// TIA Portal project "Inteligenta_szklarnia" (V15.1)

(* hardware
DEVICE "S7-1200 station_2"  S7-1200 Station
   slot 0: "Rack_0"  S7-1200 Rack  Rack  V1.0
   slot 1: "PLC_1"  CPU 1214C AC/DC/Rly  6ES7 214-1BE30-0XB0  V2.2
DEVICE "HMI_1"  KTP700 Basic PN
   slot 0: "HMI_1"  KTP700 Basic PN  6AV2 123-2GB03-0AX0  15.1.0.0
   slot 1: "HMI_RT_3"  KTP700 Basic PN  6AV2 123-2GB03-0AX0  15.1.0.0
   slot 5: "HMI_1.IE_CP_1"  PROFINET Interface  15.0.1.0
      slot 1: "PROFINET Interface_1"  PROFINET Interface
         slot 1: "Port_1"  Port
DEVICE "S7-1200 station_1"  S7-1200 Station
   slot 0: "Rack_0"  S7-1200 Rack  Rack  V1.0
   slot 1: "PLC_do_symulacji"  CPU 1214C AC/DC/Rly  6ES7 214-1BG40-0XB0  V4.2
DEVICE "HMI_do_symulacji"  KTP700 Basic PN
   slot 0: "HMI_do_symulacji"  KTP700 Basic PN  6AV2 123-2GB03-0AX0  15.1.0.0
   slot 1: "HMI_RT_2"  KTP700 Basic PN  6AV2 123-2GB03-0AX0  15.1.0.0
   slot 5: "HMI_do_symulacji.IE_CP_1"  PROFINET Interface  15.0.1.0
      slot 1: "PROFINET Interface_1"  PROFINET Interface
         slot 1: "Port_1"  Port
*)

// ===== PLC "PLC_1"  CPU 1214C AC/DC/Rly =====

VAR_GLOBAL   // PLC tag table "Default tag table"
   "Tag_1" AT %I0.0 : Bool;
   "Tag_ScreenNumber" AT %MD0 : DInt;
   "FirstScan" AT %M1.0 : Bool;
   "DiagStatusUpdate" AT %M1.1 : Bool;
   "AlwaysTRUE" AT %M1.2 : Bool;
   "AlwaysFALSE" AT %M1.3 : Bool;
END_VAR

VAR_GLOBAL   // PLC tag table "wyjscia"
   "Grzałka" AT %Q0.0 : Bool;
   "Wentylator" AT %Q0.1 : Bool;
   "Pompa_wodna" AT %Q0.2 : Bool;
   "Rolety_zamykanie" AT %Q0.4 : Bool;
   "Alarm_ostrzegwaczy" AT %Q0.5 : Bool;
   "Siłownik_okien_otwieranie" AT %Q0.6 : Bool;
   "Siłownik_okien_zamykanie" AT %Q0.7 : Bool;
   "Rolety_otwieranie" AT %Q0.3 : Bool;
END_VAR

DATA_BLOCK "Parametry"   // DB1
{ S7_Optimized_Access := 'TRUE' }
VERSION : 0.1
   VAR
      Wilgotność_powietrza : Int;
      Wilgotność_gleby : Int;
      temeratura : Real;
      Czujnik_światła : Int;
      Czujnik_wiatru : Int;
      czujnik_CO2 : Int;
      stopien_zasloniecia_rolet : Int;
   END_VAR
BEGIN
END_DATA_BLOCK

DATA_BLOCK "Wejscia_HMI"   // DB2
{ S7_Optimized_Access := 'TRUE' }
VERSION : 0.1
   VAR
      Temperatura : Real;
      CO2 : Real;
      Wilgotność_gleby : Int;
      Wilgotność_powietrza : Int;
      Zaciemnienie : Int;
      naslonecznienie_manual : Int;
   END_VAR
BEGIN
END_DATA_BLOCK

DATA_BLOCK "Receptury"   // DB3
{ S7_Optimized_Access := 'TRUE' }
VERSION : 0.1
   VAR
      nasłonecznienie : Array[0..5] of Int;
      system_okien : Array[0..5] of Bool;
      wilgotnosc_gleby : Array[0..5] of Int;
      wilgotnosc_powietrza : Array[0..5] of Int;
      temperatua : Array[0..5] of Real;
      nazwa : Array[0..5] of String;
   END_VAR
BEGIN
END_DATA_BLOCK

DATA_BLOCK "Archiwizowane_parametry"   // DB4
{ S7_Optimized_Access := 'TRUE' }
VERSION : 0.1
   VAR
      Temperatura : Array[0..335] of Real;
      Wilgotnosc : Array[0..335] of Int;
      Naslonecznienie : Array[0..335] of Int;
      iterator : Int := 0;   // Iterator służący do zapisu danych w odpowiednich komórkach tablicy.
      Zerowanie : Array[0..335] of Int;
   END_VAR
BEGIN
   Naslonecznienie[0] := 0;
   Naslonecznienie[1] := 0;
END_DATA_BLOCK

// folder: System blocks/Program resources

DATA_BLOCK "IEC_Timer_0_DB"   // DB5
{ S7_Optimized_Access := 'TRUE' }
AUTHOR : Simatic
FAMILY : IEC
NAME : IEC_TMR
VERSION : 1.0
// stored: InstanceOfName IEC_TIMER
"IEC_TIMER"
BEGIN
END_DATA_BLOCK

// folder: (top level)

FUNCTION "Rolety" : Void   // FC1, LAD
{ S7_Optimized_Access := 'TRUE' }
VERSION : 0.1
   VAR_INPUT
      Czy_automatyczny : Bool;
      Czy_manualny : Bool;
   END_VAR
   VAR_TEMP   // added for the SCL form of the ladder/FBD networks
      _w1 : Bool;
   END_VAR
BEGIN

REGION Network 1: Sterowanie roletami w trybie automatycznym
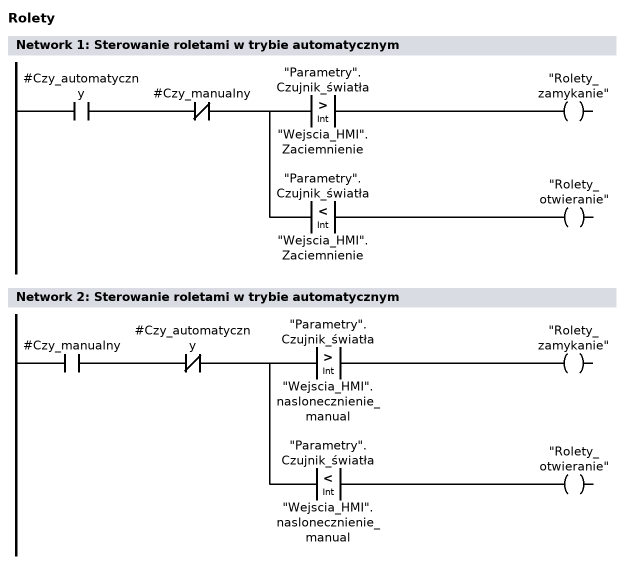
   RUNG wire#powerrail
      Contact( #Czy_automatyczny )
      I_Contact( #Czy_manualny )
      wire#w1
      { S7_Templates := "SrcType := Int" } GT_Contact(in1 := "Parametry".Czujnik_światła, in2 := "Wejscia_HMI".Zaciemnienie)
      Coil( "Rolety_zamykanie" )
   END_RUNG
   RUNG wire#w1
      { S7_Templates := "SrcType := Int" } LT_Contact(in1 := "Parametry".Czujnik_światła, in2 := "Wejscia_HMI".Zaciemnienie)
      Coil( "Rolety_otwieranie" )
   END_RUNG
   // the same network as SCL:
   #_w1 := #Czy_automatyczny AND NOT #Czy_manualny;
   "Rolety_zamykanie" := #_w1 AND ("Parametry".Czujnik_światła > "Wejscia_HMI".Zaciemnienie);
   "Rolety_otwieranie" := #_w1 AND ("Parametry".Czujnik_światła < "Wejscia_HMI".Zaciemnienie);
END_REGION

REGION Network 2: Sterowanie roletami w trybie automatycznym
   RUNG wire#powerrail
      Contact( #Czy_manualny )
      I_Contact( #Czy_automatyczny )
      wire#w1
      { S7_Templates := "SrcType := Int" } GT_Contact(in1 := "Parametry".Czujnik_światła, in2 := "Wejscia_HMI".naslonecznienie_manual)
      Coil( "Rolety_zamykanie" )
   END_RUNG
   RUNG wire#w1
      { S7_Templates := "SrcType := Int" } LT_Contact(in1 := "Parametry".Czujnik_światła, in2 := "Wejscia_HMI".naslonecznienie_manual)
      Coil( "Rolety_otwieranie" )
   END_RUNG
   // the same network as SCL:
   #_w1 := #Czy_manualny AND NOT #Czy_automatyczny;
   "Rolety_zamykanie" := #_w1 AND ("Parametry".Czujnik_światła > "Wejscia_HMI".naslonecznienie_manual);
   "Rolety_otwieranie" := #_w1 AND ("Parametry".Czujnik_światła < "Wejscia_HMI".naslonecznienie_manual);
END_REGION
END_FUNCTION

FUNCTION "Archiwizacja_parametrow" : Void   // FC2, LAD
{ S7_Optimized_Access := 'TRUE' }
VERSION : 0.1
// Zapis parametrów do bloku DB odbywa się co pół godziny. Po uruchomieniu sterownika pierwszy zapis nie odbywa się od razu, aby wykres nie przedstawiał parametrów, które nie były jeszcze regulowane.
BEGIN

REGION Network 1
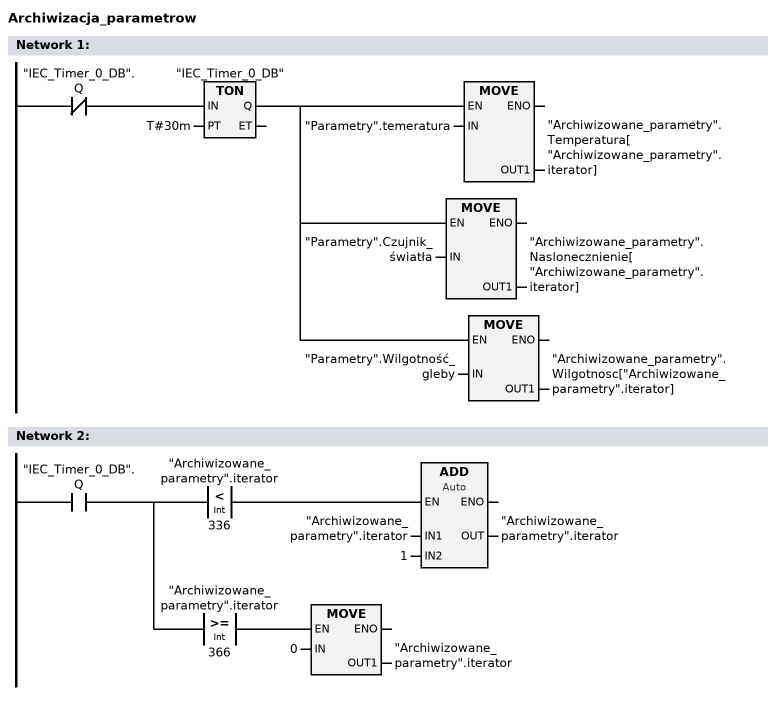
   "IEC_Timer_0_DB".TON(IN := NOT "IEC_Timer_0_DB".Q, PT := T#30m);
   IF "IEC_Timer_0_DB".Q THEN
       "Archiwizowane_parametry".Temperatura["Archiwizowane_parametry".iterator] := "Parametry".temeratura;
       "Archiwizowane_parametry".Naslonecznienie["Archiwizowane_parametry".iterator] := "Parametry".Czujnik_światła;
       "Archiwizowane_parametry".Wilgotnosc["Archiwizowane_parametry".iterator] := "Parametry".Wilgotność_gleby;
   END_IF;
END_REGION

REGION Network 2
   RUNG wire#powerrail
      Contact( "IEC_Timer_0_DB".Q )
      wire#w1
      { S7_Templates := "SrcType := Int" } LT_Contact(in1 := "Archiwizowane_parametry".iterator, in2 := 336)
      { S7_GenerateENO := "TRUE" } Add(in1 := "Archiwizowane_parametry".iterator, in2 := 1, out => "Archiwizowane_parametry".iterator)
   END_RUNG
   RUNG wire#w1
      { S7_Templates := "SrcType := Int" } GE_Contact(in1 := "Archiwizowane_parametry".iterator, in2 := 366)
      { S7_GenerateENO := "TRUE" } Move(in := 0, out1 => "Archiwizowane_parametry".iterator)
   END_RUNG
   // the same network as SCL:
   IF "IEC_Timer_0_DB".Q AND ("Archiwizowane_parametry".iterator < 336) THEN
       "Archiwizowane_parametry".iterator := "Archiwizowane_parametry".iterator + 1;
   END_IF;
   IF "IEC_Timer_0_DB".Q AND ("Archiwizowane_parametry".iterator >= 366) THEN
       "Archiwizowane_parametry".iterator := 0;
   END_IF;
END_REGION
END_FUNCTION

ORGANIZATION_BLOCK "Main"   // OB1, LAD, ProgramCycle
TITLE = "Main Program Sweep (Cycle)"
{ S7_Optimized_Access := 'TRUE' }
VERSION : 0.1
   VAR_INPUT
      Initial_Call : Bool;   // Initial call of this OB
      Remanence : Bool;   // =True, if remanent data are available
   END_VAR
BEGIN

REGION Network 1
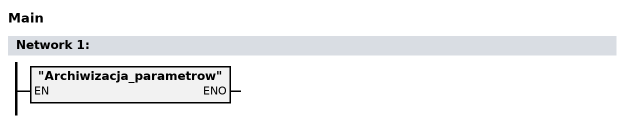
   RUNG wire#powerrail
      "Archiwizacja_parametrow"()
   END_RUNG
   // the same network as SCL:
   "Archiwizacja_parametrow"();
END_REGION
END_ORGANIZATION_BLOCK

ORGANIZATION_BLOCK "Startup"   // OB100, LAD, Startup
TITLE = "Complete Restart"
{ S7_Optimized_Access := 'TRUE' }
VERSION : 0.1
   VAR_INPUT
      LostRetentive : Bool;   // True if retentive data are lost
      LostRTC : Bool;   // True if date and time are lost
   END_VAR
BEGIN

REGION Network 1
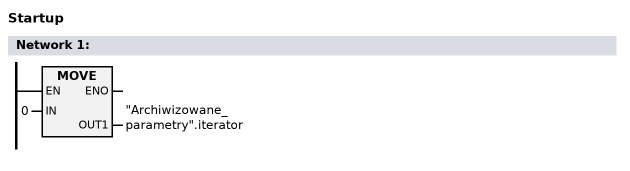
   RUNG wire#powerrail
      { S7_GenerateENO := "TRUE" } Move(in := 0, out1 => "Archiwizowane_parametry".iterator)
   END_RUNG
   // the same network as SCL:
   "Archiwizowane_parametry".iterator := 0;
END_REGION
END_ORGANIZATION_BLOCK

// ===== PLC "PLC_do_symulacji"  CPU 1214C AC/DC/Rly =====

VAR_GLOBAL   // PLC tag table "Default tag table"
   "Tag_1" AT %M0.0 : Bool;
   "System_Byte" AT %MB1 : Byte;
   "FirstScan" AT %M1.0 : Bool;
   "DiagStatusUpdate" AT %M1.1 : Bool;
   "AlwaysTRUE" AT %M1.2 : Bool;
   "AlwaysFALSE" AT %M1.3 : Bool;
   "Tag_2" AT %M0.1 : Bool;
   "Clock_Byte" AT %MB30 : Byte;
   "Clock_10Hz" AT %M30.0 : Bool;
   "Clock_5Hz" AT %M30.1 : Bool;
   "Clock_2.5Hz" AT %M30.2 : Bool;
   "Clock_2Hz" AT %M30.3 : Bool;
   "Clock_1.25Hz" AT %M30.4 : Bool;
   "Clock_1Hz" AT %M30.5 : Bool;
   "Clock_0.625Hz" AT %M30.6 : Bool;
   "Clock_0.5Hz" AT %M30.7 : Bool;
END_VAR

VAR_GLOBAL   // PLC tag table "wyjscia"
   "Grzałka" AT %Q0.0 : Bool;
   "Wentylator" AT %Q0.1 : Bool;
   "Pompa_zraszacze" AT %Q0.2 : Bool;   // Pompa zraszaczy, które odpowiadają za wilgotność powietrza w szklarni
   "Rolety_zamykanie" AT %Q0.4 : Bool;
   "Alarm_ostrzegwaczy" AT %Q0.5 : Bool;
   "Siłownik_okien_otwieranie" AT %Q0.6 : Bool;
   "Siłownik_okien_zamykanie" AT %Q0.7 : Bool;
   "Rolety_otwieranie" AT %Q0.3 : Bool;
   "Pompa_podlewanie" AT %Q1.0 : Bool;   // Pompa podlewania kropelkowego, która odpowiada za wilgotność gleby
END_VAR

DATA_BLOCK "Wejscia_PLC"   // DB1
{ S7_Optimized_Access := 'TRUE' }
VERSION : 0.1
   VAR
      Czujnik_wilgotności_powietrza : Int;   // Czujnik wilgotności powietrza w szklarni
      Czujnik_wilgotności_gleby : Int;   // Czujnik wilgotności gleby w szklarni
      Temperatura_wewnetrzna : Real;   // Temperatura wewnątrz szklarni
      Czujnik_natezenia_swiatła : Int;   // Czujnik natężenia światła wewnątrz szklarni
      Czujnik_wiatru : Int;   // Czujnik prędkości wiatru poza szklarnią
      Wewnetrzny_czujnik_CO2 : Int;   // Czujnik stężenia dwutlenku węgla w szklarni
      Stopien_zasloniecia_rolet : Int;   // Stopień zasłonięcia rolet w szklarni (przyjęty przedział 0-100%)
      Temperatura_zewnetrzna : Real;   // Temperatura mierzona na zewnątrz, poza szklarnią. Typ Int, ponieważ nie jest wymagana taka dokładność jak w pomiarze temperatury wewnętrznej.
      Zewnetrzny_czujnik_CO2 : Int;   // Czujnik stężenia dwutlenku węgla poza szklarnią
      czujnik_wilgotnosci_zewnetrzny : Int := 50;   // Potrzebny w ramach symulacji realnych warunkow
   END_VAR
BEGIN
END_DATA_BLOCK

DATA_BLOCK "HMI"   // DB2
{ S7_Optimized_Access := 'TRUE' }
VERSION : 0.1
   VAR
      nazwa_receptury : String;
      System_okien_auto : Bool;   // Wł/wył system okien w trybie automatycznym
      Przycisk_zraszacze_manual : Bool;   // Przycisk pompy zraszaczy w trybie manualnym
      Przycisk_podlewanie_manual : Bool;   // Przycisk pompy podlewania w trybie manualnym
      Przycisk_grzanie_manual : Bool;   // Przycisk grzałki w trybie manualnym
      Przycisk_wentylacja_manual : Bool;   // Przycisk wentylacji w trybie manualnym
      Otwarcie_okien_manual : Bool;   // Ustawiony w trybie manualnym otwarcie okien
      Stopien_zasloniecia_rolet_manual : Int;   // Ustawiony w trybie manualnym stopień zasłonięcia rolet
      Temperatura_auto : Real := 22.0;   // Nastawiona temeratura w trybie automatycznym
      Naslonecznienie_auto : Int := 1000;   // Nastawiona wartość nasłonecznienia w trybie automatycznym
      Wilgotnosc_powietrza_auto : Int := 50;   // Nastawiona wartość wilgotności powietrza w trybie automatycznym
      Poziom_CO2_auto : Int := 800;   // Nastawiona wartość stężenia CO2 w trybie automatycznym
      Wilgotnosc_gleby_auto : Int := 60;   // Nastawiona wartość wilgotności gleby w trybie automatycznym
      Przycisk_zatwierdz_auto : Bool;   // Przycisk zatwierdzający wcześniej wybrane ustawienia trybu automatycznego
      Przycisk_zatwierdz_zapis_receptury : Bool;   // Przycisk zatwierdzający wcześniej wybrane ustawienia trybu zapisania receptury
      Przycisk_zatwierdz_wybor_receptury : Bool;   // Przycisk zatwierdzający wcześniej wybrane ustawienia trybu receptury
      Numer_ekranu_HMI : Int;   // Numer aktualnie otwartego ekranu w HMI
      Aktywacja_trybu_manualnego : Bool;
      Aktywacja_trybu_automatycznego : Bool;
      Aktywacja_trybu_Receptur : Bool;
      Aktywacja_trybu_zapis_Receptur : Bool;
   END_VAR
BEGIN
END_DATA_BLOCK

DATA_BLOCK "Tryb_auto_parametry"   // DB7
{ S7_Optimized_Access := 'TRUE' }
VERSION : 0.1
   VAR
      nazwa : String;
      Temperatura : Real;
      Naslonecznienie : Int;
      Wilgotnosc_powietrza : Int;
      Wilgotnosc_gleby : Int;
      System_okien : Bool;
      Stezenie_co2 : Int;
   END_VAR
BEGIN
END_DATA_BLOCK

DATA_BLOCK "Alarmy"   // DB9
{ S7_Optimized_Access := 'TRUE' }
VERSION : 0.1
   VAR
      Warning_niska_temp : String := 'Zbyt niska wartość temperatury utrzymuje się długi czas. Sprawdź grzałkę lub czujnik temperatury.';   // Treść ostrzeżenia wyświetlającego się, gdy temperatura przez długi czas mieści się poniżej wymaganej wartości
      Warning_niska_temp_1 : Bool;
      Warning_wysoka_temp : String := 'Zbyt wysoka wartość temperatury utrzymuje się długi czas. Sprawdź wentylator lub czujnik temperatury.';   // Treść ostrzeżenia wyświetlającego się, gdy temperatura przez długi czas mieści się powyżej wymaganej wartości
      Warning_wysoka_temp_1 : Bool;
      Warning_nieprawidlowe_CO2 : String := 'Stężenie CO2 w zklarni przez długi czas nie osiąga prawidłowych wartości!';   // Treść ostrzeżenia wyświetlającego się, gdy stężenie CO2 w szklarni nie mieści się przez długi czas w wymaganym zakresie
      Warning_nieprawidlowe_CO2_1 : Bool;
      Blad_zbyt_wysokie_CO2 : String := 'Stężenie CO2 w szklarni ma zbyt wysoki poziom. Należy otworzyć okna, uruchomić wentylator lub podjąć inn działania.';   // Treść błędu wyświetlającego się, gdy stężenie CO2 w szklarni ma zbyt wysoki poziom.
      Blad_zbyt_wysokie_CO2_1 : Bool;
   END_VAR
BEGIN
END_DATA_BLOCK

// folder: Archiwizacja_parametrow

DATA_BLOCK "Archiwizowane_parametry"   // DB4
{ S7_Optimized_Access := 'TRUE' }
VERSION : 0.1
   VAR
      Temperatura : Array[0..335] of Real;
      Wilgotnosc : Array[0..335] of Int;
      Naslonecznienie : Array[0..335] of Int;
      iterator : Int := 0;   // Iterator służący do zapisu danych w odpowiednich komórkach tablicy.
   END_VAR
BEGIN
   Naslonecznienie[0] := 0;
   Naslonecznienie[1] := 0;
END_DATA_BLOCK

// folder: System blocks/Program resources

DATA_BLOCK "IEC_Timer_0_DB_4"   // DB3
{ S7_Optimized_Access := 'TRUE' }
AUTHOR : Simatic
FAMILY : IEC
NAME : IEC_TMR
VERSION : 1.0
// stored: InstanceOfName IEC_TIMER
"IEC_TIMER"
BEGIN
END_DATA_BLOCK

DATA_BLOCK "IEC_Timer_0_DB"   // DB5
{ S7_Optimized_Access := 'TRUE' }
AUTHOR : Simatic
FAMILY : IEC
NAME : IEC_TMR
VERSION : 1.0
// stored: InstanceOfName IEC_TIMER
"IEC_TIMER"
BEGIN
END_DATA_BLOCK

DATA_BLOCK "IEC_Timer_0_DB_1"   // DB6
{ S7_Optimized_Access := 'TRUE' }
AUTHOR : Simatic
FAMILY : IEC
NAME : IEC_TMR
VERSION : 1.0
// stored: InstanceOfName IEC_TIMER
"IEC_TIMER"
BEGIN
END_DATA_BLOCK

DATA_BLOCK "IEC_Timer_0_DB_2"   // DB8
{ S7_Optimized_Access := 'TRUE' }
AUTHOR : Simatic
FAMILY : IEC
NAME : IEC_TMR
VERSION : 1.0
// stored: InstanceOfName IEC_TIMER
"IEC_TIMER"
BEGIN
END_DATA_BLOCK

DATA_BLOCK "IEC_Timer_0_DB_5"   // DB10
{ S7_Optimized_Access := 'TRUE' }
AUTHOR : Simatic
FAMILY : IEC
NAME : IEC_TMR
VERSION : 1.0
// stored: InstanceOfName IEC_TIMER
"IEC_TIMER"
BEGIN
END_DATA_BLOCK

DATA_BLOCK "IEC_Timer_0_DB_3"   // DB11
{ S7_Optimized_Access := 'TRUE' }
AUTHOR : Simatic
FAMILY : IEC
NAME : IEC_TMR
VERSION : 1.0
// stored: InstanceOfName IEC_TIMER
"IEC_TIMER"
BEGIN
END_DATA_BLOCK

DATA_BLOCK "IEC_Counter_0_DB"   // DB12
{ S7_Optimized_Access := 'TRUE' }
AUTHOR : Simatic
FAMILY : IEC
NAME : CNTR
VERSION : 1.0
// stored: InstanceOfName IEC_COUNTER
"IEC_COUNTER"
BEGIN
END_DATA_BLOCK

// folder: (top level)

FUNCTION "Rolety" : Void   // FC1, LAD
{ S7_Optimized_Access := 'TRUE' }
VERSION : 0.1
   VAR_INPUT
      Czy_automatyczny : Bool;
      Czy_manualny : Bool;
   END_VAR
BEGIN

REGION Network 1: Warunki otwierania rolet w trybie automatycznym i manualnym
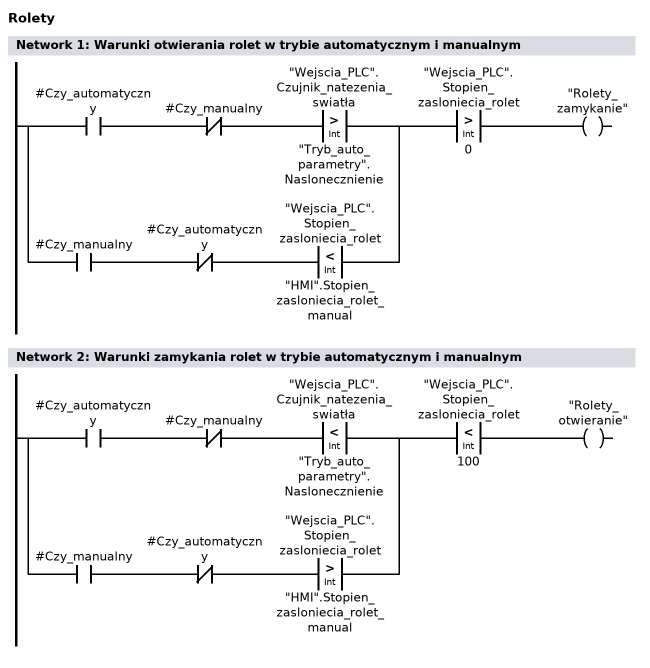
   RUNG wire#powerrail
      Contact( #Czy_automatyczny )
      I_Contact( #Czy_manualny )
      { S7_Templates := "SrcType := Int" } GT_Contact(in1 := "Wejscia_PLC".Czujnik_natezenia_swiatła, in2 := "Tryb_auto_parametry".Naslonecznienie)
      wire#w1
      { S7_Templates := "SrcType := Int" } GT_Contact(in1 := "Wejscia_PLC".Stopien_zasloniecia_rolet, in2 := 0)
      Coil( "Rolety_zamykanie" )
   END_RUNG
   RUNG wire#powerrail
      Contact( #Czy_manualny )
      I_Contact( #Czy_automatyczny )
      { S7_Templates := "SrcType := Int" } LT_Contact(in1 := "Wejscia_PLC".Stopien_zasloniecia_rolet, in2 := "HMI".Stopien_zasloniecia_rolet_manual)
   END_RUNG wire#w1
   // the same network as SCL:
   "Rolety_zamykanie" := ((#Czy_automatyczny AND NOT #Czy_manualny AND ("Wejscia_PLC".Czujnik_natezenia_swiatła > "Tryb_auto_parametry".Naslonecznienie)) OR (#Czy_manualny AND NOT #Czy_automatyczny AND ("Wejscia_PLC".Stopien_zasloniecia_rolet < "HMI".Stopien_zasloniecia_rolet_manual))) AND ("Wejscia_PLC".Stopien_zasloniecia_rolet > 0);
END_REGION

REGION Network 2: Warunki zamykania rolet w trybie automatycznym i manualnym
   RUNG wire#powerrail
      Contact( #Czy_automatyczny )
      I_Contact( #Czy_manualny )
      { S7_Templates := "SrcType := Int" } LT_Contact(in1 := "Wejscia_PLC".Czujnik_natezenia_swiatła, in2 := "Tryb_auto_parametry".Naslonecznienie)
      wire#w1
      { S7_Templates := "SrcType := Int" } LT_Contact(in1 := "Wejscia_PLC".Stopien_zasloniecia_rolet, in2 := 100)
      Coil( "Rolety_otwieranie" )
   END_RUNG
   RUNG wire#powerrail
      Contact( #Czy_manualny )
      I_Contact( #Czy_automatyczny )
      { S7_Templates := "SrcType := Int" } GT_Contact(in1 := "Wejscia_PLC".Stopien_zasloniecia_rolet, in2 := "HMI".Stopien_zasloniecia_rolet_manual)
   END_RUNG wire#w1
   // the same network as SCL:
   "Rolety_otwieranie" := ((#Czy_automatyczny AND NOT #Czy_manualny AND ("Wejscia_PLC".Czujnik_natezenia_swiatła < "Tryb_auto_parametry".Naslonecznienie)) OR (#Czy_manualny AND NOT #Czy_automatyczny AND ("Wejscia_PLC".Stopien_zasloniecia_rolet > "HMI".Stopien_zasloniecia_rolet_manual))) AND ("Wejscia_PLC".Stopien_zasloniecia_rolet < 100);
END_REGION
END_FUNCTION

FUNCTION "Sterowanie_grzalka_wentylator" : Void   // FC3, LAD
{ S7_Optimized_Access := 'TRUE' }
VERSION : 0.1
   VAR_INPUT
      czy_manualny : Bool;
      czy_automatyczny : Bool;
   END_VAR
   VAR_TEMP
      Histereza_minus : Real;   // Wartość zadanej temperatury zmieniona o dolną wartość hiterezy
      Histereza_plus : Real;   // Wartość zadanej temperatury zmieniona o górną wartość hiterezy
   END_VAR
   VAR CONSTANT
      Wartosc_histerezy : Real := 1.0;
   END_VAR
   VAR_TEMP   // added for the SCL form of the ladder/FBD networks
      _w1 : Bool;
   END_VAR
BEGIN

REGION Network 1: Sterowanie wentylatorem w trybie automatycznym i manualnym
   // Gdy uruchomiony jest tryb automatyczny, wartość temperatury w szklarni powinna się mieścić w zakresie temperatury nastawionej +- wartość histerezy. Gdy jest ona za wysoka uruchamiany jest wentylator. W trybie manualnym włączany jest on od razu po naciśnięciu przycisku do niego przypisanego.
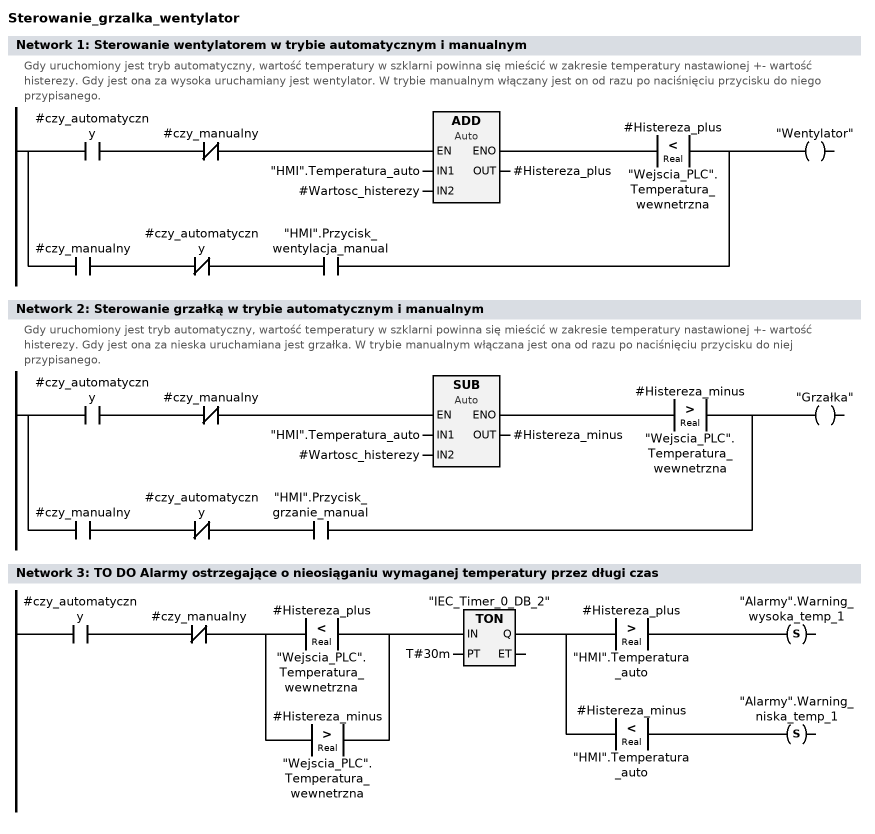
   RUNG wire#powerrail
      Contact( #czy_automatyczny )
      I_Contact( #czy_manualny )
      Add(in1 := "HMI".Temperatura_auto, in2 := #Wartosc_histerezy, out => #Histereza_plus)
      { S7_Templates := "SrcType := Real" } LT_Contact(in1 := #Histereza_plus, in2 := "Wejscia_PLC".Temperatura_wewnetrzna)
      wire#w1
      Coil( "Wentylator" )
   END_RUNG
   RUNG wire#powerrail
      Contact( #czy_manualny )
      I_Contact( #czy_automatyczny )
      Contact( "HMI".Przycisk_wentylacja_manual )
   END_RUNG wire#w1
   // the same network as SCL:
   #_w1 := #czy_automatyczny AND NOT #czy_manualny;
   IF #_w1 THEN #Histereza_plus := "HMI".Temperatura_auto + #Wartosc_histerezy; END_IF;
   "Wentylator" := (#_w1 AND (#Histereza_plus < "Wejscia_PLC".Temperatura_wewnetrzna)) OR (#czy_manualny AND NOT #czy_automatyczny AND "HMI".Przycisk_wentylacja_manual);
END_REGION

REGION Network 2: Sterowanie grzałką w trybie automatycznym i manualnym
   // Gdy uruchomiony jest tryb automatyczny, wartość temperatury w szklarni powinna się mieścić w zakresie temperatury nastawionej +- wartość histerezy. Gdy jest ona za nieska uruchamiana jest grzałka. W trybie manualnym włączana jest ona od razu po naciśnięciu przycisku do niej przypisanego.
   RUNG wire#powerrail
      Contact( #czy_automatyczny )
      I_Contact( #czy_manualny )
      Sub(in1 := "HMI".Temperatura_auto, in2 := #Wartosc_histerezy, out => #Histereza_minus)
      { S7_Templates := "SrcType := Real" } GT_Contact(in1 := #Histereza_minus, in2 := "Wejscia_PLC".Temperatura_wewnetrzna)
      wire#w1
      Coil( "Grzałka" )
   END_RUNG
   RUNG wire#powerrail
      Contact( #czy_manualny )
      I_Contact( #czy_automatyczny )
      Contact( "HMI".Przycisk_grzanie_manual )
   END_RUNG wire#w1
   // the same network as SCL:
   #_w1 := #czy_automatyczny AND NOT #czy_manualny;
   IF #_w1 THEN #Histereza_minus := "HMI".Temperatura_auto - #Wartosc_histerezy; END_IF;
   "Grzałka" := (#_w1 AND (#Histereza_minus > "Wejscia_PLC".Temperatura_wewnetrzna)) OR (#czy_manualny AND NOT #czy_automatyczny AND "HMI".Przycisk_grzanie_manual);
END_REGION

REGION Network 3: TO DO Alarmy ostrzegające o nieosiąganiu wymaganej temperatury przez długi czas
   "IEC_Timer_0_DB_2".TON(IN := #czy_automatyczny AND NOT #czy_manualny AND ((#Histereza_plus < "Wejscia_PLC".Temperatura_wewnetrzna) OR (#Histereza_minus > "Wejscia_PLC".Temperatura_wewnetrzna)),
                          PT := T#30m);
   IF "IEC_Timer_0_DB_2".Q AND (#Histereza_plus > "HMI".Temperatura_auto) THEN
       "Alarmy".Warning_wysoka_temp_1 := TRUE;
   END_IF;
   IF "IEC_Timer_0_DB_2".Q AND (#Histereza_minus < "HMI".Temperatura_auto) THEN
       "Alarmy".Warning_niska_temp_1 := TRUE;
   END_IF;
END_REGION
END_FUNCTION

FUNCTION "Zapis_parametrow_trybu_auto" : Void   // FC4, LAD
{ S7_Optimized_Access := 'TRUE' }
VERSION : 0.1
BEGIN

REGION Network 1: Zapis wybranych na HMI parametrów, aby zostały one stałe do kolejnego zatwierdzenia ich zmiany.
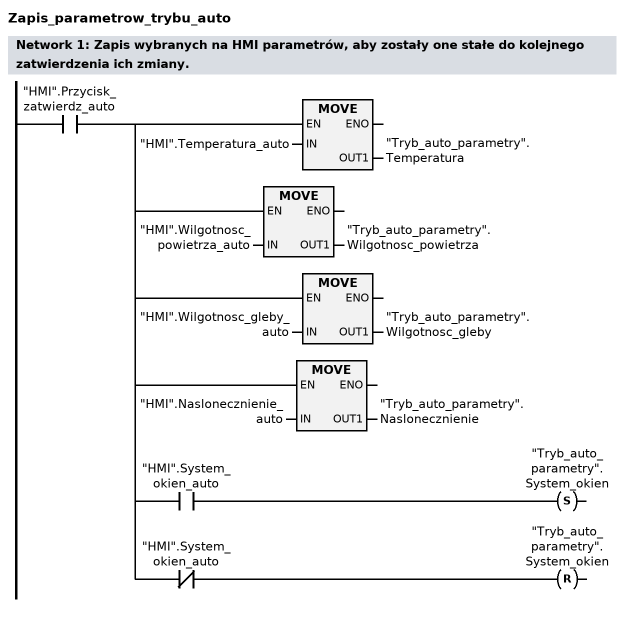
   RUNG wire#powerrail
      Contact( "HMI".Przycisk_zatwierdz_auto )
      wire#w1
      Move(in := "HMI".Temperatura_auto, out1 => "Tryb_auto_parametry".Temperatura)
   END_RUNG
   RUNG wire#w1
      Move(in := "HMI".Wilgotnosc_powietrza_auto, out1 => "Tryb_auto_parametry".Wilgotnosc_powietrza)
   END_RUNG
   RUNG wire#w1
      Move(in := "HMI".Wilgotnosc_gleby_auto, out1 => "Tryb_auto_parametry".Wilgotnosc_gleby)
   END_RUNG
   RUNG wire#w1
      Move(in := "HMI".Naslonecznienie_auto, out1 => "Tryb_auto_parametry".Naslonecznienie)
   END_RUNG
   RUNG wire#w1
      Contact( "HMI".System_okien_auto )
      S_Coil( "Tryb_auto_parametry".System_okien )
   END_RUNG
   RUNG wire#w1
      I_Contact( "HMI".System_okien_auto )
      R_Coil( "Tryb_auto_parametry".System_okien )
   END_RUNG
   // the same network as SCL:
   IF "HMI".Przycisk_zatwierdz_auto THEN
       "Tryb_auto_parametry".Temperatura := "HMI".Temperatura_auto;
       "Tryb_auto_parametry".Wilgotnosc_powietrza := "HMI".Wilgotnosc_powietrza_auto;
       "Tryb_auto_parametry".Wilgotnosc_gleby := "HMI".Wilgotnosc_gleby_auto;
       "Tryb_auto_parametry".Naslonecznienie := "HMI".Naslonecznienie_auto;
   END_IF;
   IF "HMI".Przycisk_zatwierdz_auto AND "HMI".System_okien_auto THEN
       "Tryb_auto_parametry".System_okien := TRUE;
   END_IF;
   IF "HMI".Przycisk_zatwierdz_auto AND NOT "HMI".System_okien_auto THEN
       "Tryb_auto_parametry".System_okien := FALSE;
   END_IF;
END_REGION
END_FUNCTION

FUNCTION "Jaki_Tryb" : Void   // FC5, LAD
{ S7_Optimized_Access := 'TRUE' }
VERSION : 0.1
BEGIN

REGION Network 1: Reset trybu auto jesli wykryje jakikolwiek inny tryb
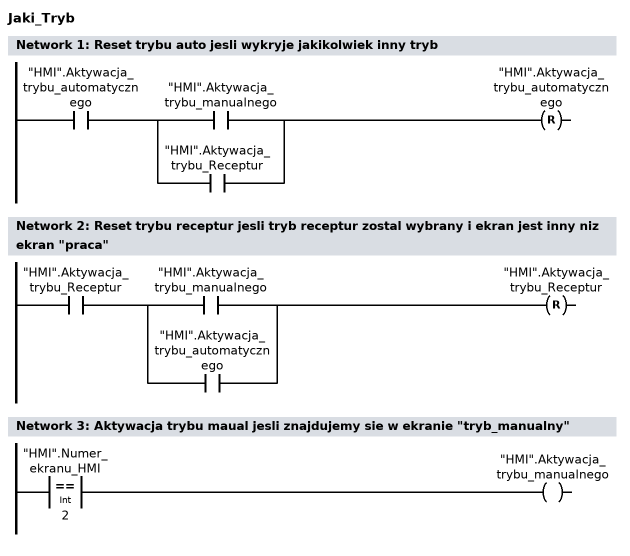
   RUNG wire#powerrail
      Contact( "HMI".Aktywacja_trybu_automatycznego )
      wire#w1
      Contact( "HMI".Aktywacja_trybu_manualnego )
      wire#w2
      R_Coil( "HMI".Aktywacja_trybu_automatycznego )
   END_RUNG
   RUNG wire#w1
      Contact( "HMI".Aktywacja_trybu_Receptur )
   END_RUNG wire#w2
   // the same network as SCL:
   IF "HMI".Aktywacja_trybu_automatycznego AND ("HMI".Aktywacja_trybu_manualnego OR "HMI".Aktywacja_trybu_Receptur) THEN
       "HMI".Aktywacja_trybu_automatycznego := FALSE;
   END_IF;
END_REGION

REGION Network 2: Reset trybu receptur jesli tryb receptur zostal wybrany i ekran jest inny niz ekran "praca"
   RUNG wire#powerrail
      Contact( "HMI".Aktywacja_trybu_Receptur )
      wire#w1
      Contact( "HMI".Aktywacja_trybu_manualnego )
      wire#w2
      R_Coil( "HMI".Aktywacja_trybu_Receptur )
   END_RUNG
   RUNG wire#w1
      Contact( "HMI".Aktywacja_trybu_automatycznego )
   END_RUNG wire#w2
   // the same network as SCL:
   IF "HMI".Aktywacja_trybu_Receptur AND ("HMI".Aktywacja_trybu_manualnego OR "HMI".Aktywacja_trybu_automatycznego) THEN
       "HMI".Aktywacja_trybu_Receptur := FALSE;
   END_IF;
END_REGION

REGION Network 3: Aktywacja trybu maual jesli znajdujemy sie w ekranie "tryb_manualny"
   RUNG wire#powerrail
      { S7_Templates := "SrcType := Int" } EQ_Contact(in1 := "HMI".Numer_ekranu_HMI, in2 := 2)
      Coil( "HMI".Aktywacja_trybu_manualnego )
   END_RUNG
   // the same network as SCL:
   "HMI".Aktywacja_trybu_manualnego := "HMI".Numer_ekranu_HMI = 2;
END_REGION
END_FUNCTION

FUNCTION "Sterowanie_podlewaniem_zraszaniem" : Void   // FC7, LAD
{ S7_Optimized_Access := 'TRUE' }
VERSION : 0.1
   VAR_INPUT
      Czy_automatyczny : Bool;
      Czy_manualny : Bool;
   END_VAR
BEGIN

REGION Network 1: Sterowanie pompą zraszaczy, które odpowiadają za wilgotność powietrza w szklarni
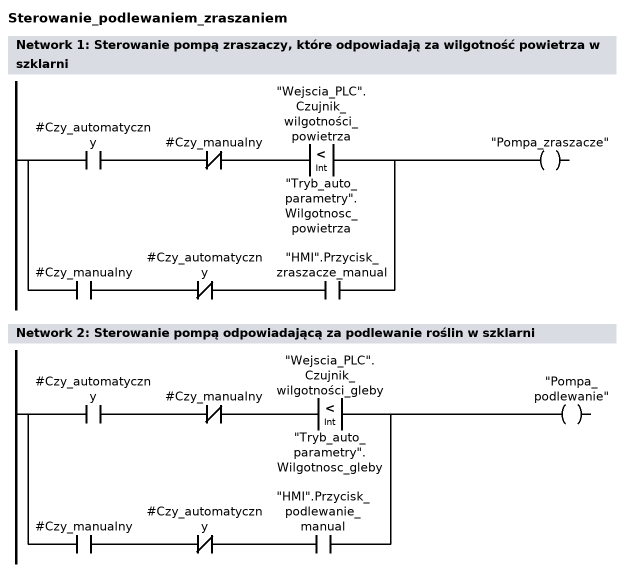
   RUNG wire#powerrail
      Contact( #Czy_automatyczny )
      I_Contact( #Czy_manualny )
      { S7_Templates := "SrcType := Int" } LT_Contact(in1 := "Wejscia_PLC".Czujnik_wilgotności_powietrza, in2 := "Tryb_auto_parametry".Wilgotnosc_powietrza)
      wire#w1
      Coil( "Pompa_zraszacze" )
   END_RUNG
   RUNG wire#powerrail
      Contact( #Czy_manualny )
      I_Contact( #Czy_automatyczny )
      Contact( "HMI".Przycisk_zraszacze_manual )
   END_RUNG wire#w1
   // the same network as SCL:
   "Pompa_zraszacze" := (#Czy_automatyczny AND NOT #Czy_manualny AND ("Wejscia_PLC".Czujnik_wilgotności_powietrza < "Tryb_auto_parametry".Wilgotnosc_powietrza)) OR (#Czy_manualny AND NOT #Czy_automatyczny AND "HMI".Przycisk_zraszacze_manual);
END_REGION

REGION Network 2: Sterowanie pompą odpowiadającą za podlewanie roślin w szklarni
   RUNG wire#powerrail
      Contact( #Czy_automatyczny )
      I_Contact( #Czy_manualny )
      { S7_Templates := "SrcType := Int" } LT_Contact(in1 := "Wejscia_PLC".Czujnik_wilgotności_gleby, in2 := "Tryb_auto_parametry".Wilgotnosc_gleby)
      wire#w1
      Coil( "Pompa_podlewanie" )
   END_RUNG
   RUNG wire#powerrail
      Contact( #Czy_manualny )
      I_Contact( #Czy_automatyczny )
      Contact( "HMI".Przycisk_podlewanie_manual )
   END_RUNG wire#w1
   // the same network as SCL:
   "Pompa_podlewanie" := (#Czy_automatyczny AND NOT #Czy_manualny AND ("Wejscia_PLC".Czujnik_wilgotności_gleby < "Tryb_auto_parametry".Wilgotnosc_gleby)) OR (#Czy_manualny AND NOT #Czy_automatyczny AND "HMI".Przycisk_podlewanie_manual);
END_REGION
END_FUNCTION

FUNCTION "Sterowanie_oknami" : Void   // FC8, LAD
{ S7_Optimized_Access := 'TRUE' }
VERSION : 0.1
   VAR_INPUT
      czy_manualny : Bool;
      czy_automatyczny : Bool;
   END_VAR
   VAR_TEMP
      Histereza_plus : Int;
      Histereza_minus : Int;
      Zakres_temp_gora : Real;   // Górny zakres temperatury zewnętrznej dla której w trybie automatycznym będą otwierane okna
      Zakres_temp_dol : Real;   // Dolny zakres temperatury zewnętrznej dla której w trybie automatycznym będą otwierane okna
   END_VAR
   VAR CONSTANT
      Histereza : Int := 25;   // Histereza, która określa kiedy stan CO2 w szklarni jest uznawany za prawidłowy
   END_VAR
BEGIN

REGION Network 1: Operacje matematyczne używane w networku 2. i 3.
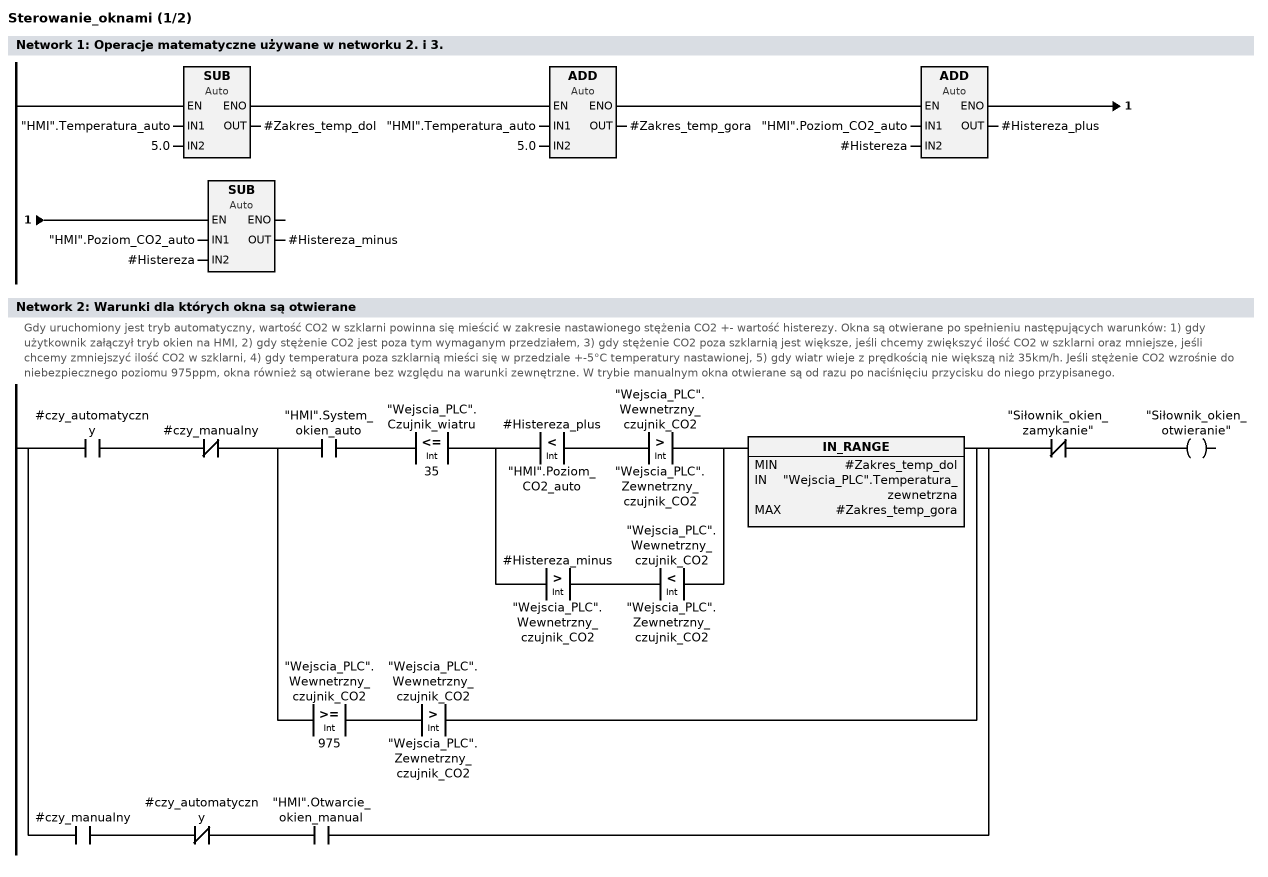
   RUNG wire#powerrail
      Sub(in1 := "HMI".Temperatura_auto, in2 := 5.0, out => #Zakres_temp_dol)
      Add(in1 := "HMI".Temperatura_auto, in2 := 5.0, out => #Zakres_temp_gora)
      Add(in1 := "HMI".Poziom_CO2_auto, in2 := #Histereza, out => #Histereza_plus)
      Sub(in1 := "HMI".Poziom_CO2_auto, in2 := #Histereza, out => #Histereza_minus)
   END_RUNG
   // the same network as SCL:
   #Zakres_temp_dol := "HMI".Temperatura_auto - 5.0;
   #Zakres_temp_gora := "HMI".Temperatura_auto + 5.0;
   #Histereza_plus := "HMI".Poziom_CO2_auto + #Histereza;
   #Histereza_minus := "HMI".Poziom_CO2_auto - #Histereza;
END_REGION
